VERSION : 1.1
// The FC checks if a given token is a parameter
   VAR_INPUT
      tokenToCheck : Struct   // struct of actual and previous token to be checked
         actual : String;   // actual token
         previous : String;   // previous token
      END_STRUCT;
      language : Int;   // language package selection
      lastIndexLookUp : DInt;   // last index in lookUpTable
   END_VAR
   VAR_IN_OUT
      parameterDefinition : "LKinLang_typeParameterDefinition";   // parameter definiton
      parameterLookUpTable : Array[1.."LKINLANG_MAX_NUMBER_OF_PARAMETERS"] of "LKinLang_typeParameterLookUp";   // lookUpTable for given language
      parameterDefaults : Variant;   // default parameter values
      directCmdWord : Word;   // word for direct command
      configCmdWords : Array[1.."LKINLANG_NUMBER_OF_FOLLOW_VALUES"] of Word;   // words for configuration commands
   END_VAR
   VAR_TEMP
      tempCounter : Int;   // temporary counter variable
      tempSeparator : Array[1.."LKINLANG_NUMBER_OF_SEPARATORS"] of Byte;   // temporary variable for separators array
      tempMerger : Array[1.."LKINLANG_NUMBER_OF_MERGERS"] of Byte;   // temporary variable for mergers array
      tempValidCounts : "LKinLang_typePathDataElementCounter";   // temporary variable for valid counts
      tempParameterNameNumber : DInt;   // temporary variable for parameter name number
      tempString : "LKinLang_typeVariableDeclaration";
      tempKeyToken : "LKinLang_typeKeyToken";
   END_VAR
   // Ret_Val : parameter assigned to token
BEGIN
   //==========================================================================================
   // SIEMENS AG
   // (c)Copyright 2019 All Rights Reserved
   //------------------------------------------------------------------------------------------
   // Library: LKinLang
   // Tested with: S7-1517T-3 PN/DP
   // Engineering: TIA Portal V15
   // Restrictions: ---
   // Requirements: S7-1500T FW 2.5
   // Functionality: LKinLang_IsTokenParameter
   // The FC checks if a given token is a parameter
   // 
   // Support: tech.team.motioncontrol@siemens.com
   // Note: Parameter comments are only available in language 'English (United States)'
   //------------------------------------------------------------------------------------------
   // Change log table:
   // Version    Date          Expert in charge    Changes applied
   // 01.00.00   28.05.2019    FR                  First created version
   //===========================================================================================

   //======================================================================
   // Is token a known parameter - return: parameter number for array
   //======================================================================
   // Check parameters with parameter number (>-1)
   // Initialize --> no match
   #LKinLang_IsTokenParameter := 0;

   IF "LKinLang_IsTokenNumberInclSign"(#tokenToCheck.previous) THEN
     #tempParameterNameNumber := STRING_TO_DINT(#tokenToCheck.previous);
   ELSE
     #tempParameterNameNumber := -1;
   END_IF;


   // Search in array for string with number
   FOR #tempCounter := 1 TO #lastIndexLookUp DO
     IF #parameterLookUpTable[#tempCounter].parameterNameString = #tokenToCheck.actual
       AND (#parameterLookUpTable[#tempCounter].parameterNameNumber = #tempParameterNameNumber
       OR #parameterLookUpTable[#tempCounter].parameterNameNumber = -1)
     THEN

       // Get definition
       "LKinLang_SelectLangPackage"(language := #language,
                                    variableDeclarations=>#tempString,
                                    keyToken=>#tempKeyToken,
                                    parameterDefinition := #parameterDefinition,
                                    separators => #tempSeparator,
                                    mergers => #tempMerger,
                                    validCounts => #tempValidCounts,
                                    parameterNumber := #parameterLookUpTable[#tempCounter].parameterNumber,
                                    parameterDefaults := #parameterDefaults);


       #directCmdWord := #parameterLookUpTable[#tempCounter].directValueWord;
       #configCmdWords := #parameterLookUpTable[#tempCounter].followValueWords;

       #LKinLang_IsTokenParameter := DINT_TO_USINT(#parameterLookUpTable[#tempCounter].parameterNumber);
       RETURN;
     ELSE
       ;
     END_IF;
   END_FOR;
END_FUNCTION

FUNCTION "LKinLang_IsTokenSeparator" : USInt   // FC35473, SCL
TITLE = LKinLang_IsTokenSeparator
{ S7_Optimized_Access := 'TRUE' }
AUTHOR : tech.team.motioncontrol@siemens.com
FAMILY : LKinLang
VERSION : 1.1
// The FC checks if a given token is a separator
   VAR_IN_OUT
      tokenToCheck : String;   // token to be checked
      separators : Array[1.."LKINLANG_NUMBER_OF_SEPARATORS"] of Byte;   // array of separators
   END_VAR
   VAR_TEMP
      tempSeparatorIndex : Int;   // temporary variable storing separator index in string
   END_VAR
   // Ret_Val : parameter assigned to separator token
BEGIN
   //==========================================================================================
   // SIEMENS AG
   // (c)Copyright 2019 All Rights Reserved
   //------------------------------------------------------------------------------------------
   // Library: LKinLang
   // Tested with: S7-1517T-3 PN/DP
   // Engineering: TIA Portal V15
   // Restrictions: ---
   // Requirements: S7-1500T FW 2.5
   // Functionality: LKinLang_IsTokenSeparator
   // The FC checks if a given token is a separator
   // 
   // Support: tech.team.motioncontrol@siemens.com
   // Note: Parameter comments are only available in language 'English (United States)'
   //------------------------------------------------------------------------------------------
   // Change log table:
   // Version    Date          Expert in charge    Changes applied
   // 01.00.00   28.05.2019    FR                  First created version
   //===========================================================================================

   //======================================================================
   // Is token a known parameter - return: parameter number for array
   //======================================================================

   // Initialize variables
   #LKinLang_IsTokenSeparator := 0;
   #tempSeparatorIndex := 0;

   // Check if token is one single separator    
   IF LEN(#tokenToCheck) = 1 THEN

     //Check for separator
     //--------------------------------------------------------------------------------
     // compare sign with all separators
     FOR #tempSeparatorIndex := 1 TO "LKINLANG_NUMBER_OF_SEPARATORS" DO
       // detect separator
       IF #separators[#tempSeparatorIndex] = #tokenToCheck[1] THEN
         // Set separator index
         #LKinLang_IsTokenSeparator := INT_TO_USINT(#tempSeparatorIndex);
         EXIT;
       ELSE
         ; // no match
       END_IF;

     END_FOR;
   ELSE
     // more than one sign -> can´t be a single separator
     #LKinLang_IsTokenSeparator := 0;
   END_IF;
END_FUNCTION

FUNCTION "LKinLang_IsTokenVariable" : Void   // FC35474, SCL
TITLE = LKinLang_IsTokenVariable
{ S7_Optimized_Access := 'TRUE' }
AUTHOR : tech.team.motioncontrol@siemens.com
FAMILY : LKinLang
VERSION : 1.0
// The FC checks if a given token is a variable
   VAR_INPUT
      lineNumber : UDInt;   // Line number
      tokenCheck : Struct   // Struct with the token to check
         actual : String;
         previous : String;
      END_STRUCT;
   END_VAR
   VAR_OUTPUT
      varIndex : Int;   // Variable index
      varType : Int;   // Varaible type
   END_VAR
   VAR_IN_OUT
      varRefList : "LKinLang_typeVarRefList";   // Variables reference list
      keyToken : "LKinLang_typeKeyToken";   // Key token to find variables
      subPrgList : "LKinLang_typeSubPrgList";   // Subprogram list
      errorString : String;   // Error string connection
      stringExpression : String;   // String expression
   END_VAR
   VAR_TEMP
      tempCounter : DInt;   // Temporary counter
      tempMaxIndex : Int;   // Temporary max index
      tempCurrentScope : DInt;   // Temporary scope
   END_VAR
BEGIN
   //==========================================================================================
   // SIEMENS AG
   // (c)Copyright 2020 All Rights Reserved
   //------------------------------------------------------------------------------------------
   // Library: LKinLang
   // Tested with: S7-1517T-3 PN/DP
   // Engineering: TIA Portal V15
   // Restrictions: ---
   // Requirements: S7-1500T FW 2.5
   // Functionality: LKinLang_IsTokenVariable
   // The FC checks if a given token is a variable
   // 
   // Support: tech.team.motioncontrol@siemens.com
   // Note: Parameter comments are only available in language 'English (United States)'
   //------------------------------------------------------------------------------------------
   // Change log table:
   // Version    Date          Expert in charge    Changes applied
   // 01.00.00   24.11.2020    FR                  First created version
   //===========================================================================================

   //======================================================================
   // Is token (or any other string) a variable
   //======================================================================
   // Check if it is an interface variable
   // Line look like this:
   // X = %I8
   // 
   // Token:
   // [1] 8
   // [2] %I
   // [3] 
   // [4] =
   // [5] 
   // [6] X
   // 
   // OR
   //
   // Token:
   // [1] 1000
   // [2] =
   // [3] 1
   // [4] %I
   // 

   // Init outputs
   #varType := 0;
   #varIndex := 0;

   // Define current scope 
   IF #subPrgList.subPrgs[1].lineNumberStart = 0 // If no sub exists the scope is also set to 1
       OR #lineNumber < #subPrgList.subPrgs[1].lineNumberStart
   THEN
       #tempCurrentScope := 1;
   ELSE
       FOR #tempCounter := 1 TO #subPrgList.numberOfSubPrgs DO
           IF #lineNumber > #subPrgList.subPrgs[#tempCounter].lineNumberStart
               AND #lineNumber < #subPrgList.subPrgs[#tempCounter].lineNumberEnd
           THEN
               #tempCurrentScope := 10 * #tempCounter;
           ELSE
               CONTINUE;
           END_IF;
       END_FOR;
   END_IF;


   IF #tokenCheck.actual = #keyToken.tokenInterfaceVarBool THEN
       // Set the var type to Bool 
       #varType := "LKINLANG_VAR_TYPE_INTERFACE_BOOL";
   ELSIF #tokenCheck.actual = #keyToken.tokenInterfaceVarDInt THEN
       // Set the var type to DInt
       #varType := "LKINLANG_VAR_TYPE_INTERFACE_DINT";
   ELSIF #tokenCheck.actual = #keyToken.tokenInterfaceVarLReal THEN
       // Set the var type to LReal
       #varType := "LKINLANG_VAR_TYPE_INTERFACE_LREAL";
   ELSE
       // Check if token is a local variable
       // Count backwards --> Local should be found before global
       FOR #tempCounter := #varRefList.numberOfReferences TO 1 BY -1 DO
           // Check if actual token is a variable name in the ref table
           IF #tokenCheck.actual = #varRefList.references[#tempCounter].name THEN
               // Check if scope is matching
               IF #tempCurrentScope = #varRefList.references[#tempCounter].scope
                   OR #varRefList.references[#tempCounter].scope = 2 // Global scope
               THEN
                   // Token is variable
                   // Get name, type and index
                   #varIndex := #varRefList.references[#tempCounter].index;
                   #varType := #varRefList.references[#tempCounter].type;
                   #errorString := '';
                   EXIT;
               ELSE
                   // error --> scope is not valid
                   #errorString := '';
                   #errorString := CONCAT(IN1 := #errorString, IN2 := 'Error: Cannot access variable out of scope');
                   #errorString := CONCAT(IN1 := #errorString, IN2 := ' in line: ');
                   #errorString := CONCAT(IN1 := #errorString, IN2 := UDINT_TO_STRING(#lineNumber));
                   CONTINUE; // Continue searching if name is duplicate, scope could match later
               END_IF;
           END_IF;
       END_FOR;
   END_IF;

   // Token is any kind of interface variable 
   IF #varType >= "LKINLANG_VAR_TYPE_INTERFACE_BOOL" THEN
     // the index should be the previous token
     IF "LKinLang_IsTokenNumberInclSign"(#tokenCheck.previous) THEN
       #varIndex := STRING_TO_INT(#tokenCheck.previous);
       // Remove index from stringExpression
       #stringExpression := RIGHT(IN := #stringExpression,
                                  L := LEN(#stringExpression) - LEN(#tokenCheck.previous));
     ELSE
       // error --> index is not a number
       #errorString := CONCAT(IN1 := #errorString, IN2 := 'Error: Interface variable index wrong or missing');
       #errorString := CONCAT(IN1 := #errorString, IN2 := ' in line: ');
       #errorString := CONCAT(IN1 := #errorString, IN2 := UDINT_TO_STRING(#lineNumber));
     END_IF;

   END_IF;

   // Check index of variable depending on type
   CASE #varType OF
     "LKINLANG_VAR_TYPE_LOCAL_BOOL": // local bool
       #tempMaxIndex := "LKINLANG_NUMBER_OF_LOCAL_BOOL";

     "LKINLANG_VAR_TYPE_LOCAL_DINT": // local dint
       #tempMaxIndex := "LKINLANG_NUMBER_OF_LOCAL_DINT";

     "LKINLANG_VAR_TYPE_LOCAL_LREAL": // local lreal
       #tempMaxIndex := "LKINLANG_NUMBER_OF_LOCAL_LREAL";

     "LKINLANG_VAR_TYPE_INTERFACE_BOOL": // interface dint
       #tempMaxIndex := "LKINLANG_NUMBER_OF_INTERFACE_BOOL";

     "LKINLANG_VAR_TYPE_INTERFACE_DINT": // interface dint
       #tempMaxIndex := "LKINLANG_NUMBER_OF_INTERFACE_DINT";

     "LKINLANG_VAR_TYPE_INTERFACE_LREAL": // interface lreal
       #tempMaxIndex := "LKINLANG_NUMBER_OF_INTERFACE_LREAL";

     ELSE
       ; // type not defined
   END_CASE;

   // Check if index is out of bounds
   IF #tempMaxIndex <> 0 AND // Check if maxIndex was set --> Var was actually found
     (#varIndex < 1 OR #varIndex > #tempMaxIndex) // Check index against bounds
   THEN 
     // error --> index is not valid
     #errorString := CONCAT(IN1 := #errorString, IN2 := 'Error: Variable index out of bounds');
     #errorString := CONCAT(IN1 := #errorString, IN2 := ' in line: ');
     #errorString := CONCAT(IN1 := #errorString, IN2 := UDINT_TO_STRING(#lineNumber));
   END_IF;
END_FUNCTION

FUNCTION "LKinLang_LRealToReducedString" : String   // FC35475, SCL
TITLE = LKinLang_LRealToReducedString
{ S7_Optimized_Access := 'TRUE' }
AUTHOR : tech.team.motioncontrol@siemens.com
FAMILY : LKinLang
VERSION : 1.1
// The FC converts an LReal to string with a given amount of decimal places
   VAR_INPUT
      input : LReal;   // LReal value to be reduced to a string
      decimalPlaces : Int;   // number of decimal digits
   END_VAR
   VAR_TEMP
      tempCompleteString : String;   // temporary variable to store complete string
      tempCounter : Int;   // temporary counter variable
      tempNumber : LReal;   // temporary variable for storing the number to be reduced
      tempDecimal : LReal;   // temporary variable storing decimal digit
      tempDecimalZero : LReal;   // temporary variable storing decimal 0
      tempDecimalDint : DInt;   // temporary variable storing decimal DInt
      tempNumberString : String;   // temporary variable storing number string
      tempDecimalString : String;   // temporary variable storing decimal string
      tempZeroString : String;   // temporary variable storing zero string
   END_VAR
   // Ret_Val : returned string created from LReal value
BEGIN
   //==========================================================================================
   // SIEMENS AG
   // (c)Copyright 2019 All Rights Reserved
   //------------------------------------------------------------------------------------------
   // Library: LKinLang
   // Tested with: S7-1517T-3 PN/DP
   // Engineering: TIA Portal V15
   // Restrictions: ---
   // Requirements: S7-1500T FW 2.5
   // Functionality: LKinLang_LRealToReducedString
   // The FC converts an LReal to string with a given amount of decimal places
   // 
   // Support: tech.team.motioncontrol@siemens.com
   // Note: Parameter comments are only available in language 'English (United States)'
   //------------------------------------------------------------------------------------------
   // Change log table:
   // Version    Date          Expert in charge    Changes applied
   // 01.00.00   28.05.2019    FR                  First created version
   // 01.00.01   17.07.2019    FR                  Added exception when decimal places = 0
   // 01.00.02   24.03.2020    FR                  Delete '+' sign from string when >= 0.0
   //                                              Fix negative values being rounded
   // 02.00.00   27.03.2020    FR                  Rework using VAL_STRG
   // 02.00.01   18.02.2021    FR                  Fix for x.0 
   //===========================================================================================

   //======================================================================
   // Returns Lreal input as String with set digits
   //======================================================================

   VAL_STRG(IN:=#input,
            SIZE:=INT_TO_USINT(MAX_LEN(#tempCompleteString)), // Length of generated string
            PREC:=INT_TO_USINT(#decimalPlaces), // Number of decimal places
            FORMAT:=0, // Format 0 means leading '-' only, decimal fraction and '.'
            P:=1, // Start with the first character
            OUT=>#tempCompleteString);

   // delete leading spaces
   FOR #tempCounter := LEN(#tempCompleteString) TO 1 BY -1 DO
     // Find first space
     IF #tempCompleteString[#tempCounter] = ' ' THEN
       #tempCompleteString := RIGHT(IN:=#tempCompleteString, L:=LEN(#tempCompleteString) - #tempCounter);
       EXIT;
     END_IF;
   END_FOR;

   // delete zeros after last digits
   FOR #tempCounter := LEN(#tempCompleteString) TO 1 BY -1 DO
     // Leave loop if decimal point is found
     IF #tempCompleteString[#tempCounter] = '.' THEN
       EXIT;
     END_IF;

     // Find first zero
     IF #tempCompleteString[#tempCounter] <> '0' THEN
       #tempCompleteString := LEFT(IN := #tempCompleteString, L := #tempCounter);
       EXIT;
     END_IF;
   END_FOR;

   // copy out ----------------------
   #LKinLang_LRealToReducedString := #tempCompleteString;
END_FUNCTION

FUNCTION "LKinLang_PostEqualsSignWhenExpressionMandCnd" : Bool   // FC35476, SCL
TITLE = LKinLang_PostEqualsSignWhenExpressionMandCnd / LKinLang_PostEqualSignWhenExpressionMandCnd
{ S7_Optimized_Access := 'TRUE' }
AUTHOR : tech.team.motioncontrol@siemens.com
FAMILY : LKinLang
VERSION : 1.1
// The FC checks if a "=" is mandatory or not permitted
   VAR_INPUT
      stringExpression : String;   // string expression to be checked
      currentTokenNo : Int;   // number of current token
      tokenOffset : Int;   // offset to number of token
   END_VAR
   VAR_IN_OUT
      lineToken : "LKinLang_typeLineTokens";   // line token
   END_VAR
   VAR_TEMP
      tempReturnValue : Bool;   // temporary variable storing return value
      tempSignIndex : Int;   // temporary variable storing index of sign
      tempTokenIndexOffset : Int;   // temporary variable storing index offset of token
      tempReturnValue2 : Bool;   // temporary variable storing return value 2
      tempAlgebraicSignAllowed : Bool;   // temporary variable algebraic sign allowed
   END_VAR
   // Ret_Val : TRUE: equals sign as following token is required; FALSE: equals sign as following token is NOT required
   VAR CONSTANT
      SPACE : String := ' ';   // Space character
      EQUAL : String := '=';   // Equal sign character
   END_VAR
BEGIN
   //==========================================================================================
   // SIEMENS AG
   // (c)Copyright 2019 All Rights Reserved
   //------------------------------------------------------------------------------------------
   // Library: LKinLang
   // Tested with: S7-1517T-3 PN/DP
   // Engineering: TIA Portal V15
   // Restrictions: ---
   // Requirements: S7-1500T FW 2.5
   // Functionality: LKinLang_PostEqualsSignWhenExpressionMandCnd
   // The FC checks if a "=" is mandatory and if yes then check spaces
   // 
   // 
   // Support: tech.team.motioncontrol@siemens.com
   // Note: Parameter comments are only available in language 'English (United States)'
   //------------------------------------------------------------------------------------------
   // Change log table:
   // Version    Date          Expert in charge    Changes applied
   // 01.00.00   28.05.2019    FR                  First created version
   // 01.01.00   15.01.2020    FR                  Back to old code with function calls
   //===========================================================================================

   // Are the last tokens togehter a number or a string? 
   //  Check if variable was used ?
   //  --> The stringExpressioon already contains the value but the token contains the var name 
   //  --> Error when using: H100=myVar
   //  --> Check token if it is a variable and then use PostEqualSignMandCnd ?

   IF "LKinLang_IsTokenNumberInclSign"(#stringExpression) THEN
     // Number: so check for the mandatory number OR the OPTIONAL "=" sign
     #tempReturnValue := "LKinLang_PostNumberMandCnd"(algebraicSignAllowed := TRUE,
                                                      currentTokenNo := #currentTokenNo,
                                                      tokenOffset := #tokenOffset,
                                                      lineTokens := #lineToken)


     OR "LKinLang_PostEqualSignMandCnd"(currentTokenNo := #currentTokenNo,
                                        tokenOffset := #tokenOffset,
                                        lineTokens := #lineToken);
   ELSE
     // String: So check for the MANDATORY "=" sign
     #tempReturnValue := "LKinLang_PostEqualSignMandCnd"(currentTokenNo := #currentTokenNo,
                                                         tokenOffset := #tokenOffset,
                                                         lineTokens := #lineToken);
   END_IF;

   // Write return value
   #LKinLang_PostEqualsSignWhenExpressionMandCnd := #tempReturnValue;
END_FUNCTION

FUNCTION "LKinLang_PostNumberMandCnd" : Bool   // FC35477, SCL
TITLE = LKinLang_PostNumberMandCnd
{ S7_Optimized_Access := 'TRUE' }
AUTHOR : tech.team.motioncontrol@siemens.com
FAMILY : LKinLang
VERSION : 1.1
// The FC checks if following token is a valid number
   VAR_INPUT
      algebraicSignAllowed : Bool;   // algebraic sign allowed
      currentTokenNo : Int;   // number of current token
      tokenOffset : Int;   // offset to number of token
   END_VAR
   VAR_IN_OUT
      lineTokens : "LKinLang_typeLineTokens";   // line token
   END_VAR
   // Ret_Val : TRUE: number as following token is required; FALSE: number as following token is NOT required
BEGIN
   //==========================================================================================
   // SIEMENS AG
   // (c)Copyright 2019 All Rights Reserved
   //------------------------------------------------------------------------------------------
   // Library: LKinLang
   // Tested with: S7-1517T-3 PN/DP
   // Engineering: TIA Portal V15
   // Restrictions: ---
   // Requirements: S7-1500T FW 2.5
   // Functionality: LKinLang_PostNumberMandCnd
   // The FC checks if following token is a valid number
   // 
   // Support: tech.team.motioncontrol@siemens.com
   // Note: Parameter comments are only available in language 'English (United States)'
   //------------------------------------------------------------------------------------------
   // Change log table:
   // Version    Date          Expert in charge    Changes applied
   // 01.00.00   28.05.2019    FR                  First created version
   //===========================================================================================

   //======================================================================
   // A Number is mandatory after Parameter, no spaces allowed.
   // Return: yes or no
   //======================================================================

   // Not first token, because there can´t be a number before
   IF #currentTokenNo >= 2 AND (#currentTokenNo - #tokenOffset - 1) >= 1 THEN
     IF #algebraicSignAllowed AND #currentTokenNo >= 3 AND (#currentTokenNo - #tokenOffset - 2) > 0 THEN
       // Is the token befor a number? Algebraic sign ALLOWED
       IF "LKinLang_IsTokenNumberInclSign"(CONCAT(IN1 := #lineTokens.lineToken[#currentTokenNo - #tokenOffset - 1], IN2 := #lineTokens.lineToken[#currentTokenNo - #tokenOffset - 2]))
         OR "LKinLang_IsTokenNumber"(#lineTokens.lineToken[#currentTokenNo - #tokenOffset - 1])
       THEN
         #LKinLang_PostNumberMandCnd := TRUE;
       ELSE
         #LKinLang_PostNumberMandCnd := FALSE;
       END_IF;
     ELSE
       // Is the token before a number? Algebraic sign forbidden
       IF "LKinLang_IsTokenNumber"(#lineTokens.lineToken[#currentTokenNo - #tokenOffset - 1]) THEN
         #LKinLang_PostNumberMandCnd := TRUE;
       ELSE
         #LKinLang_PostNumberMandCnd := FALSE;
       END_IF;
     END_IF;
   ELSE
     #LKinLang_PostNumberMandCnd := FALSE;
   END_IF;
END_FUNCTION

FUNCTION "LKinLang_PreProcessor" : Void   // FC35478, SCL
TITLE = LKinLang_PreProcessor
{ S7_Optimized_Access := 'TRUE' }
AUTHOR : tech.team.motioncontrol@siemens.com
FAMILY : LKinLang
VERSION : 1.1
// The FC replaces parts of strings in program lines
   VAR_INPUT
      preprocessorConfig : "LKinLang_typePreProcessorReplacement";   // pre processor configuration
   END_VAR
   VAR_IN_OUT
      programLine : String;   // program line to be checked and edited by pre processor
   END_VAR
   VAR_TEMP
      tempProgramLine : String;   // temporary program line
      tempCounter : DInt;   // temporary counter
      tempIndex : DInt;   // temporary counter
      tempLengthOfSearchTerm : Int;   // temporary variable for length of search term
      tempLengthOfReplaceTerm : Int;   // temporary variable for length of replace term
      tempFirstPosOfFoundString : Int;   // temporary variable for first position of found string
      tempEmptyReplace : String;   // temporary empty replacement string
   END_VAR
BEGIN
   //==========================================================================================
   // SIEMENS AG
   // (c)Copyright 2021 All Rights Reserved
   //------------------------------------------------------------------------------------------
   // Library: LKinLang
   // Tested with: S7-1517T-3 PN/DP
   // Engineering: TIA Portal V16
   // Restrictions: ---
   // Requirements: S7-1500T FW 2.8
   // Functionality: LKinLang_PreProcessor
   // The FC replaces parts of strings in program lines
   // 
   // Support: tech.team.motioncontrol@siemens.com
   // Note: Parameter comments are only available in language 'English (United States)'
   //------------------------------------------------------------------------------------------
   // Change log table:
   // Version    Date          Expert in charge    Changes applied
   // 01.00.00   28.05.2019    FR                  First created version
   // 01.00.01   15.02.2021    FR                  Added repeat for multiple replacements in the same line
   // 01.00.02   12.04.2021    FR                  Added replacement in temp
   //===========================================================================================

   //======================================================================
   // Replacements done by pre processor
   //======================================================================  

   // Initialize temp values
   #tempCounter := 0;
   #tempLengthOfSearchTerm := 0;
   #tempLengthOfReplaceTerm := 0;
   #tempFirstPosOfFoundString := 0;
   #tempProgramLine := #programLine;

   // Searching
   FOR #tempCounter := 1 TO "LKINLANG_NUMBER_OF_REPLACEMENTS" DO
     #tempLengthOfSearchTerm := LEN(#preprocessorConfig.replacements[#tempCounter].searchTerm);
     #tempLengthOfReplaceTerm := LEN(#preprocessorConfig.replacements[#tempCounter].replaceTerm);

     IF #tempLengthOfSearchTerm > 0 THEN // Search term existing
       REPEAT // Repeat replacing until no more replacements found in this line
         #tempFirstPosOfFoundString := FIND(IN1 := #tempProgramLine, IN2 := #preprocessorConfig.replacements[#tempCounter].searchTerm);
         IF #tempFirstPosOfFoundString <> 0 THEN // String was found
           #programLine := REPLACE(IN1 := #programLine,
                                   IN2 := #preprocessorConfig.replacements[#tempCounter].replaceTerm,
                                   L := #tempLengthOfSearchTerm,
                                   P := #tempFirstPosOfFoundString);

           // Create "empty" replacement string to keep tempProgramLine and ProgramLine the same length
           #tempEmptyReplace := '';
           FOR #tempIndex := 1 TO #tempLengthOfReplaceTerm DO
             #tempEmptyReplace := CONCAT(IN1 := #tempEmptyReplace, IN2 := BYTE_TO_CHAR(16#0)); // Concat NULL chars
           END_FOR;
           // Delete already processed characters from temp string to avoid endless loop
           // Replace searched term with NULL string
           #tempProgramLine := REPLACE(IN1 := #tempProgramLine, IN2 := #tempEmptyReplace, L := #tempLengthOfSearchTerm, P := #tempFirstPosOfFoundString);

         ELSE
           ; // Search term not in code line
         END_IF;

       UNTIL #tempFirstPosOfFoundString = 0 END_REPEAT;

     ELSE
       ; // No search term
     END_IF;
   END_FOR;
END_FUNCTION

FUNCTION "LKinLang_ReplaceTapsBySpaces" : Void   // FC35479, SCL
TITLE = LKinLang_ReplaceTapsBySpaces
{ S7_Optimized_Access := 'TRUE' }
AUTHOR : tech.team.motioncontrol@siemens.com
FAMILY : LKinLang
VERSION : 1.1
// The FC replaces tabs in a given string by spaces
   VAR_IN_OUT
      codeline : String;   // string to be edited
   END_VAR
   VAR_TEMP
      tempCounter : Int;   // temporary counter variable
   END_VAR
BEGIN
   //==========================================================================================
   // SIEMENS AG
   // (c)Copyright 2019 All Rights Reserved
   //------------------------------------------------------------------------------------------
   // Library: LKinLang
   // Tested with: S7-1517T-3 PN/DP
   // Engineering: TIA Portal V15
   // Restrictions: ---
   // Requirements: S7-1500T FW 2.5
   // Functionality: LKinLang_ReplaceTabsBySpaces
   // The FC replaces tabs in a given string by spaces
   // 
   // Support: tech.team.motioncontrol@siemens.com
   // Note: Parameter comments are only available in language 'English (United States)'
   //------------------------------------------------------------------------------------------
   // Change log table:
   // Version    Date          Expert in charge    Changes applied
   // 01.00.00   28.05.2019    FR                  First created version
   //===========================================================================================

   //======================================================================
   // Replace Tap ($T) and ascii zero in referenced ascii line by spaces
   //======================================================================  

   // Search tap
   FOR #tempCounter := 1 TO LEN(#codeline) DO
     IF #codeline[#tempCounter] = '$09' //16#09
       OR #codeline[#tempCounter] = '$00' //16#00
     THEN
       #codeline[#tempCounter] := '$20'; //16#20; // Replace tap trough space
     ELSE
       ; // No tap
     END_IF;
   END_FOR;
END_FUNCTION

FUNCTION "LKinLang_SetParameterConditions" : Void   // FC35480, SCL
TITLE = LKinLang_SetParameterConditions
{ S7_Optimized_Access := 'TRUE' }
AUTHOR : tech.team.motioncontrol@siemens.com
FAMILY : LKinLang
VERSION : 1.1
// The FC sets parameter conditions for given parameter numbers and definitons
   VAR_INPUT
      parameterNumber : Int;   // parameter number to be set
      tempParameterDef : "LKinLang_typeParameterDefinition";   // parameter definition for given parameter number
   END_VAR
   VAR_IN_OUT
      parametersInLine : Array[1.."LKINLANG_NUMBER_OF_CONDITIONS"] of "LKinLang_typeCondition";   // parameters programmed in actual line
      parametersInCommand : Array[1.."LKINLANG_NUMBER_OF_CONDITIONS"] of "LKinLang_typeCondition";   // parameters programmed in actual command
      parametersInProgram : Array[1.."LKINLANG_NUMBER_OF_CONDITIONS"] of "LKinLang_typeCondition";   // parameters programmed in actual program
      conditionsToCheck : Array[1.."LKINLANG_NUMBER_OF_CONDITIONS"] of "LKinLang_typeCondition";   // conditions from parameters which are to be checked
      conditionCounter : Int;   // counter for conditions array
   END_VAR
   VAR_TEMP
      tempCounter : Int;   // temporary counter variable
   END_VAR
BEGIN
   //==========================================================================================
   // SIEMENS AG
   // (c)Copyright 2019 All Rights Reserved
   //------------------------------------------------------------------------------------------
   // Library: LKinLang
   // Tested with: S7-1517T-3 PN/DP
   // Engineering: TIA Portal V15
   // Restrictions: ---
   // Requirements: S7-1500T FW 2.5
   // Functionality: LKinLang_SetParameterConditions
   // The FC sets parameter conditions for given parameter numbers and definitons
   // 
   // Support: tech.team.motioncontrol@siemens.com
   // Note: Parameter comments are only available in language 'English (United States)'
   //------------------------------------------------------------------------------------------
   // Change log table:
   // Version    Date          Expert in charge    Changes applied
   // 01.00.00   28.05.2019    FR                  First created version
   //===========================================================================================

   // Write set parameters into arrays (line/command/program)
   // Write conditions to be checked from parameter into array

   // TODO: Overflow check 

   // Write into condition array
   IF #parameterNumber <> 0 THEN

     // Conditions in line
     FOR #tempCounter := 1 TO "LKINLANG_NUMBER_OF_CONDITIONS" DO
       IF #parametersInLine[#tempCounter].ParameterNumber = #parameterNumber THEN
         // Already in array 
         EXIT;
       END_IF;
       IF #parametersInLine[#tempCounter].ParameterNumber = 0 THEN
         #parametersInLine[#tempCounter].ParameterNumber := #parameterNumber;
         EXIT;
       END_IF;
     END_FOR;

    // Command conditions  
     FOR #tempCounter := 1 TO "LKINLANG_NUMBER_OF_CONDITIONS" DO
       IF #parametersInCommand[#tempCounter].ParameterNumber = #parameterNumber THEN
         // Already in array 
         EXIT;
       END_IF;
       IF #parametersInCommand[#tempCounter].ParameterNumber = 0 THEN
         #parametersInCommand[#tempCounter].ParameterNumber := #parameterNumber;
         EXIT;
       END_IF;
     END_FOR;

     // Program conditions
     FOR #tempCounter := 1 TO "LKINLANG_NUMBER_OF_CONDITIONS" DO
       IF #parametersInProgram[#tempCounter].ParameterNumber = #parameterNumber THEN
         // Already in array 
         EXIT;
       END_IF;
       IF #parametersInProgram[#tempCounter].ParameterNumber = 0 THEN
         #parametersInProgram[#tempCounter].ParameterNumber := #parameterNumber;
         EXIT;
       END_IF;
     END_FOR;

     // Write into condition array which conditions have to be checked
     FOR #tempCounter := 1 TO "LKINLANG_NUMBER_OF_CONDITIONS" DO
       IF #tempParameterDef.conditions[#tempCounter].Group <> 0 THEN
         #conditionsToCheck[#conditionCounter] := #tempParameterDef.conditions[#tempCounter];
         #conditionCounter += 1;
       ELSE
         RETURN; // Return if group = 0 --> no more conditions follow
       END_IF;
     END_FOR;
   END_IF;
END_FUNCTION

FUNCTION "LKinLang_PostEqualSignMandCnd" : Bool   // FC35481, SCL
TITLE = LKinLang_PostEqualSignMandCnd
{ S7_Optimized_Access := 'TRUE' }
AUTHOR : tech.team.motioncontrol@siemens.com
FAMILY : LKinLang
VERSION : 1.1
// Check for mandatory '=' after condition
   VAR_INPUT
      lineTokens : "LKinLang_typeLineTokens";   // line token
      currentTokenNo : Int;   // number of current token
      tokenOffset : Int;   // offset to number of token
   END_VAR
   VAR_TEMP
      tempTokenIndexOffset : Int;   // Temporary counter to iterate through tokens
      tempTokenOffset : Int;   // Temporary offset to the token counter
   END_VAR
   // Ret_Val : TRUE: correct syntax; FALSE: wrong syntax
   VAR CONSTANT
      SPACE : Char := ' ';   // Space character
      EQUAL : Char := '=';   // Equal sign character
   END_VAR
BEGIN
   //==========================================================================================
   // SIEMENS AG
   // (c)Copyright 2020 All Rights Reserved
   //------------------------------------------------------------------------------------------
   // Library: LKinLang
   // Tested with: S7-1517T-3 PN/DP
   // Engineering: TIA Portal V15
   // Restrictions: ---
   // Requirements: S7-1500T FW 2.5
   // Functionality: LKinLang_PostEqualSignMandCnd
   // The FC checks for the correct syntax when using a expression 
   // --> mandatory '=' after parameter
   // 
   // Support: tech.team.motioncontrol@siemens.com
   // Note: Parameter comments are only available in language 'English (United States)'
   //------------------------------------------------------------------------------------------
   // Change log table:
   // Version    Date          Expert in charge    Changes applied
   // 01.00.00   13.01.2020    FR                  First created version
   //===========================================================================================
   //======================================================================
   // "=" is mandatory; spaces allowed - return: yes or no
   //======================================================================

   #tempTokenIndexOffset := 1;

   // If token offset is greater 0 then reduce it by one 
   // Usually the token offset points to the next number and not the equal sign 
   // --> Reduce offset by one to check the equals sign
   // Example:
   // H100=myVar 
   // Token:
   // [4]H
   // [3]100
   // [2]=
   // [1]myVar
   //
   // --> currentTokenNo = 4
   // --> tokenOffset = 2
   // --> tempTokenIndexOffset = 1
   // --> Previous token is checked so 'myVar' is checked to be equal which is always false!
   // --> Reduce tokenOffset by 1 to check token before 'myVar'

   IF #tokenOffset > 0 THEN
     #tempTokenOffset := #tokenOffset - 1;
   ELSE
     #tempTokenOffset := #tokenOffset;
   END_IF;

   // equal sign possible ?
   IF #currentTokenNo - #tempTokenOffset > 1 THEN
     // Check if previous token is a space or '='
     IF #lineTokens.lineToken[#currentTokenNo - #tempTokenOffset - #tempTokenIndexOffset] <> #SPACE
       AND #lineTokens.lineToken[#currentTokenNo - #tempTokenOffset - #tempTokenIndexOffset] <> #EQUAL
     THEN
       //Error: next sign no space or =
       #LKinLang_PostEqualSignMandCnd := FALSE;
     ELSE
       // Increment token index if next sign isn´t a equals sign
       IF #lineTokens.lineToken[#currentTokenNo - #tempTokenOffset - #tempTokenIndexOffset] <> #EQUAL THEN
         #tempTokenIndexOffset := #tempTokenIndexOffset + 1;
       END_IF;

       // Check last option for equal sign
       IF #lineTokens.lineToken[#currentTokenNo - #tempTokenOffset - #tempTokenIndexOffset] <> #EQUAL THEN
         //Error
         #LKinLang_PostEqualSignMandCnd := FALSE;
       ELSE
         #LKinLang_PostEqualSignMandCnd := TRUE;
       END_IF;
     END_IF;
   ELSE
     // There can´t be an equals sign
     #LKinLang_PostEqualSignMandCnd := FALSE;
   END_IF;
END_FUNCTION

FUNCTION "LKinLang_SetValue" : DWord   // FC35482, SCL
TITLE = LKinLang_SetValue
{ S7_Optimized_Access := 'TRUE' }
AUTHOR : tech.team.motioncontrol@siemens.com
FAMILY : LKinLang
VERSION : 1.1
// The FC sets the parameter value considering priority and modality of parameters
   VAR_INPUT
      parameterValue : LReal;   // value of parameter
      parameterPriority : Int;   // priority of parameter
      validCountOfParameter : Int;   // count of valid parameter uses
      parameterValueMin : LReal;   // minimum parameter value
      parameterValueMax : LReal;   // maximum parameter value
      properties : DWord;   // properties of parameter
   END_VAR
   VAR_OUTPUT
      errorString : String;   // error information (textual)
   END_VAR
   VAR_IN_OUT
      parameterCounter : Int;   // parameter counter
      priorityCounter : Int;   // priority counter
      modalCMDPrio : Int;   // priority of command modality
      modalPRGPrio : Int;   // priority of program modality
      parameterCounterInLine : Int;   // in line parameter counter
      pathDataValue : "LKinLang_typeDiffElementaryDatatypes";   // value of PathData
      modalCMDPathDataValue : "LKinLang_typeDiffElementaryDatatypes";   // value of PathData modal command
      modalPRGPathDataValue : "LKinLang_typeDiffElementaryDatatypes";   // value of PathData modal program
   END_VAR
   VAR_TEMP
      tempSymbolName : WString;   // temporary variable storing symbol name
      tempSymbolNameLength : Int;   // temporary variable storing symbol name length
      tempParaName : String;   // temporary variable storing parameter name
      tempCounter : Int;   // temporary counter variable
      tempReturnVal : DWord;   // temporary variable storing return value
      tempDataTypes : "LKinLang_typeDiffElementaryDatatypes";   // temporary variable storing data type defaults
   END_VAR
   // Ret_Val : Return value of FC
   VAR CONSTANT
      ERR_PARAMETER_COUNTER : DWord := 16#8001;   // Error due to parameter counter too high
      ERR_PARAMETER_OVERFLOW : DWord := 16#8002;   // Error due to parameter limits exceeded
      ERR_ALREADY_SET : DWord := 16#8003;   // Error deu to parameter being already set
   END_VAR
BEGIN
   //==========================================================================================
   // SIEMENS AG
   // (c)Copyright 2019 All Rights Reserved
   //------------------------------------------------------------------------------------------
   // Library: LKinLang
   // Tested with: S7-1517T-3 PN/DP
   // Engineering: TIA Portal V15
   // Restrictions: ---
   // Requirements: S7-1500T FW 2.5
   // Functionality: LKinLang_SetValue
   // The FC sets the parameter value considering priority and modality of parameters
   // 
   // Support: tech.team.motioncontrol@siemens.com
   // Note: Parameter comments are only available in language 'English (United States)'
   //------------------------------------------------------------------------------------------
   // Change log table:
   // Version    Date          Expert in charge    Changes applied
   // 01.00.00   28.05.2019    FR                  First created version
   //===========================================================================================

   //======================================================================
   // Sets PathData values which are given directly at 'parameterValue'
   //======================================================================
   // Init 
   #LKinLang_SetValue := 16#0;
   #errorString := '';

   // Assign input value to temp
   #tempDataTypes.valueLReal := #parameterValue;

   // Count how often Parameter is in set in Command // Testing only count if cmd modal 11.12.2018
   IF #parameterPriority > "LKINLANG_PRIO_DEFAULT" AND "LKinLang_CheckProperty"(properties:=#properties, propertyToCheck := "LKINLANG_CMD_MODAL") THEN // Only count parameters when certain prio is set (2 in this case)
     #parameterCounter += 1;
   ELSIF #parameterPriority > "LKINLANG_PRIO_DEFAULT" THEN // Only count parameters when certain prio is set (greater default in this case)
     #parameterCounterInLine += 1;
   END_IF;

   // // Count how often Parameter is in set in line // Testing only count if cmd modal 11.12.2018
   // IF #parameterPriority > 2 THEN // Only count parameters when certain prio is set (2 in this case)
   //   #parameterCounterInLine += 1;
   // END_IF;

   // Check Counter
   REGION CHECK_COUNTER
     IF #parameterCounter + #parameterCounterInLine > #validCountOfParameter THEN
       // Error: ParameterCounter too high

       #LKinLang_SetValue := #ERR_PARAMETER_COUNTER;
       #tempSymbolName := GetSymbolName(variable := #parameterCounter, size := 254);
       #tempSymbolNameLength := LEN(#tempSymbolName);

       FOR #tempCounter := #tempSymbolNameLength TO 1 BY -1 DO
         IF #tempSymbolName[#tempCounter] = WChar#'.' THEN
           #tempParaName := RIGHT(IN := WSTRING_TO_STRING(#tempSymbolName), L := #tempSymbolNameLength - #tempCounter);
           EXIT;
         END_IF;
       END_FOR;

       #errorString := CONCAT(IN1 := #errorString, IN2 := ';Error: Parameter counter: ');
       #errorString := CONCAT(IN1 := #errorString, IN2 := #tempParaName);
       #errorString := CONCAT(IN1 := #errorString, IN2 := '=');
       #errorString := CONCAT(IN1 := #errorString, IN2 := INT_TO_STRING(#parameterCounter + #parameterCounterInLine));
       #errorString := CONCAT(IN1 := #errorString, IN2 := '; Allowed=');
       #errorString := CONCAT(IN1 := #errorString, IN2 := INT_TO_STRING(#validCountOfParameter));
       RETURN;
     END_IF;
   END_REGION CHECK_COUNTER

   // Check Value Limits
   REGION CHECK_LIMITS
     IF "LKinLang_CheckProperty"(properties:=#properties, propertyToCheck := "LKINLANG_CHECK_LIMITS") THEN
       #tempReturnVal := "LKinLang_CheckLimits"(parameterMinVal := #parameterValueMin,
                                            parameterMaxVal := #parameterValueMax,
                                            parameterValue := #tempDataTypes);
       IF #tempReturnVal <> 0 THEN
         // Error
         // Error: Value outside limits  
         #LKinLang_SetValue := #ERR_PARAMETER_OVERFLOW;
         #tempSymbolName := GetSymbolName(variable := #parameterCounter, size := 254);
         #tempSymbolNameLength := LEN(#tempSymbolName);

         FOR #tempCounter := #tempSymbolNameLength TO 1 BY -1 DO
           IF #tempSymbolName[#tempCounter] = WChar#'.' THEN
             #tempParaName := RIGHT(IN := WSTRING_TO_STRING(#tempSymbolName), L := #tempSymbolNameLength - #tempCounter);
             EXIT;
           END_IF;
         END_FOR;

         #errorString := CONCAT(IN1 := #errorString, IN2 := ';Error: Parameter outside limits: ');
         #errorString := CONCAT(IN1 := #errorString, IN2 := #tempParaName);
         #errorString := CONCAT(IN1 := #errorString, IN2 := '=');
         #errorString := CONCAT(IN1 := #errorString, IN2 := "LKinLang_LRealToReducedString"(input := #tempDataTypes.valueLReal, decimalPlaces := 2));
         #errorString := CONCAT(IN1 := #errorString, IN2 := '; Allowed=');
         #errorString := CONCAT(IN1 := #errorString, IN2 := "LKinLang_LRealToReducedString"(input := #parameterValueMin, decimalPlaces := 2));
         #errorString := CONCAT(IN1 := #errorString, IN2 := ';');
         #errorString := CONCAT(IN1 := #errorString, IN2 := "LKinLang_LRealToReducedString"(input := #parameterValueMax, decimalPlaces := 2));
         RETURN;
       END_IF;
     ELSE // Do not check Value limits
       #tempDataTypes.valueReal := LREAL_TO_REAL(#tempDataTypes.valueLReal);
       #tempDataTypes.valueDint := LREAL_TO_DINT(#tempDataTypes.valueLReal);
       #tempDataTypes.valueInt := LREAL_TO_INT(#tempDataTypes.valueLReal);
     END_IF;
   END_REGION CHECK_LIMITS


   // Check Priority
   REGION CHECK_PRIORITY
     IF #parameterPriority > #priorityCounter THEN // Check Priority

       // Prio is ok --> Set Value
       #priorityCounter := #parameterPriority;
       #pathDataValue := #tempDataTypes;

       // Check if program modal value has to be set (is set when prio is higher or same)
       IF "LKinLang_CheckProperty"(properties:=#properties, propertyToCheck := "LKINLANG_PRG_MODAL") AND #parameterPriority >= #modalPRGPrio THEN
         #modalPRGPathDataValue := #pathDataValue;
         #modalPRGPrio := #parameterPriority;
       END_IF;

       // Check if command modal value has to be set (is set when prio is higher)
       IF "LKinLang_CheckProperty"(properties:=#properties, propertyToCheck := "LKINLANG_CMD_MODAL") AND #parameterPriority > #modalCMDPrio THEN
         #modalCMDPathDataValue := #pathDataValue;
         #modalCMDPrio := #parameterPriority;
       END_IF;

     ELSIF #priorityCounter > "LKINLANG_PRIO_DEFAULT" AND #parameterCounter + #parameterCounterInLine > 1 THEN // Value is not default and was set once
       // Prio too low
       // Error ?
       #LKinLang_SetValue := #ERR_ALREADY_SET; //???

       #tempSymbolName := GetSymbolName(variable := #parameterCounter, size := 254);
       #tempSymbolNameLength := LEN(#tempSymbolName);

       FOR #tempCounter := #tempSymbolNameLength TO 1 BY -1 DO
         IF #tempSymbolName[#tempCounter] = WChar#'.' THEN
           #tempParaName := RIGHT(IN := WSTRING_TO_STRING(#tempSymbolName), L := #tempSymbolNameLength - #tempCounter);
           EXIT;
         END_IF;
       END_FOR;

       #errorString := CONCAT(IN1 := #errorString, IN2 := #tempParaName);
       #errorString := CONCAT(IN1 := #errorString, IN2 := ' already set with higher Priority');
       RETURN;
     ELSE
       ; // Value is default but was overwritten by other command ? 
     END_IF;
   END_REGION CHECK_PRIORITY
END_FUNCTION

